(* Logix 5000 project; controller FV vendor 1 type 14 code 217 rev 31.11; software revision 31.00; part 23 of 63 *)
(* tags used below, declared in another part *)
   CheckTimeMask : INT;
   Delphi_Does_Eng_Func : BOOL;
   FR_N255 : INT[265];   // CHECKWORDS
   FR_VB4_AV04 : PlantItem;   // VB4_AV04
   FR_VB4_AV05 : PlantItem;   // VB4_AV05
   FR_VB4_AV06 : PlantItem;   // VB4_AV06
   FR_VB4_AV07 : PlantItem;   // VB4_AV07
   FR_VB4_AV08 : PlantItem;   // VB4_AV08
   FR_VB4_AV09 : PlantItem;   // VB4_AV09
   FR_VB4_AV10 : PlantItem;   // VB4_AV10
   FR_VB4_AV11 : PlantItem;   // VB4_AV11
   FR_VB4_AV12 : PlantItem;   // VB4_AV12
   FR_VB4_AV13 : PlantItem;   // VB4_AV13
   FR_VB4_AV14 : PlantItem;   // VB4_AV14
   FR_VB4_AV15 : PlantItem;   // VB4_AV15
   FR_VB4_AV23 : PlantItem;   // VB4_AV23
   TempChecktime : DINT;
(* FR_Common, continued *)

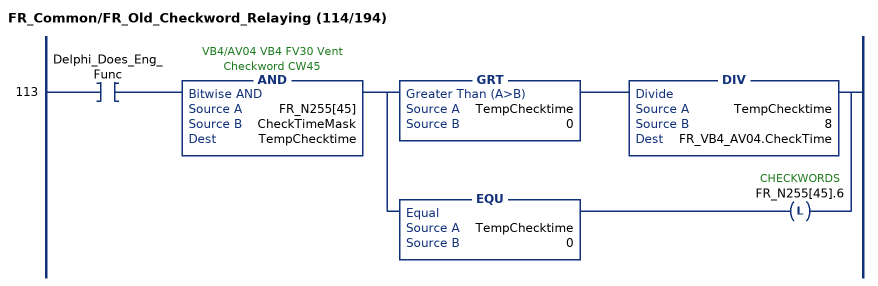
   [picture p418: FR_Common/FR_Old_Checkword_Relaying rungs 113-113]
   113: XIC(Delphi_Does_Eng_Func)AND(FR_N255[45],CheckTimeMask,TempChecktime)[GRT(TempChecktime,0) DIV(TempChecktime,8,FR_VB4_AV04.CheckTime) ,EQU(TempChecktime,0) OTL(FR_N255[45].6) ];
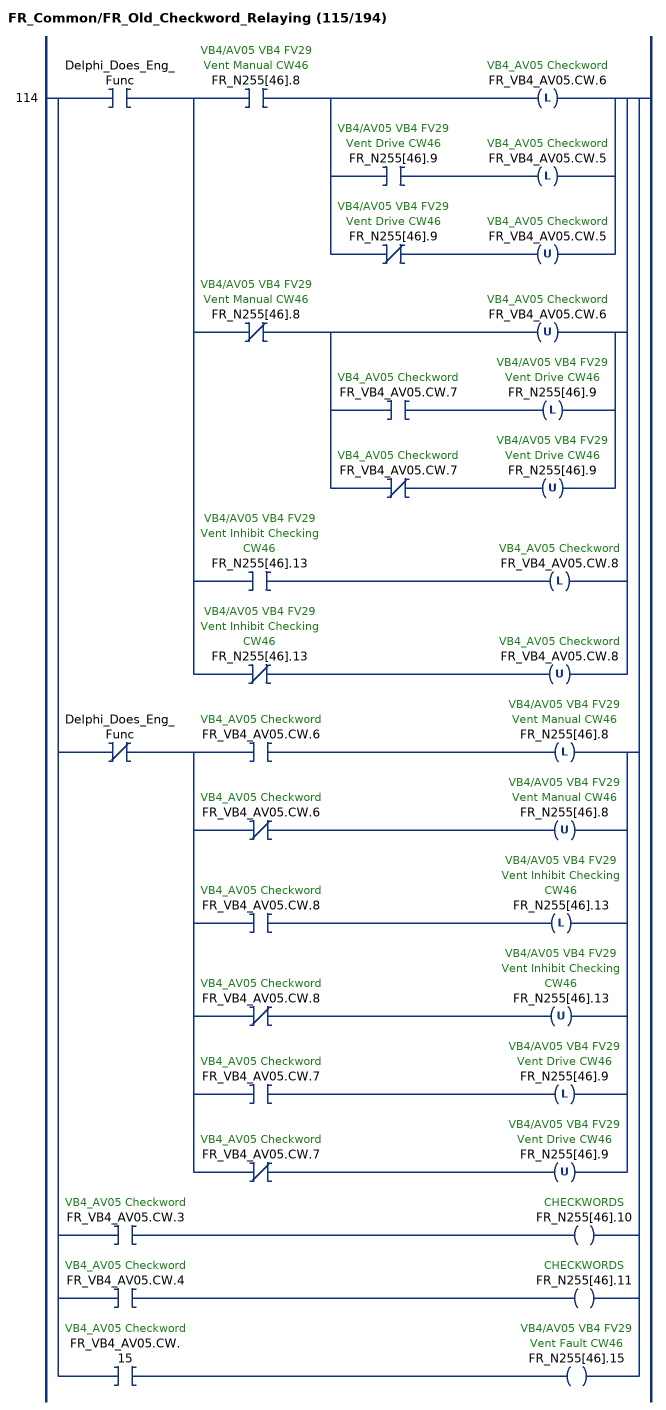
   114: [XIC(Delphi_Does_Eng_Func) [[XIC(FR_N255[46].8) [OTL(FR_VB4_AV05.CW.6) ,XIC(FR_N255[46].9) OTL(FR_VB4_AV05.CW.5) ,XIO(FR_N255[46].9) OTU(FR_VB4_AV05.CW.5) ] ,XIO(FR_N255[46].8) [OTU(FR_VB4_AV05.CW.6) ,[XIC(FR_VB4_AV05.CW.7) OTL(FR_N255[46].9) ,XIO(FR_VB4_AV05.CW.7) OTU(FR_N255[46].9) ] ] ] ,[XIC(FR_N255[46].13) OTL(FR_VB4_AV05.CW.8) ,XIO(FR_N255[46].13) OTU(FR_VB4_AV05.CW.8) ] ] ,XIO(Delphi_Does_Eng_Func) [[XIC(FR_VB4_AV05.CW.6) OTL(FR_N255[46].8) ,XIO(FR_VB4_AV05.CW.6) OTU(FR_N255[46].8) ] ,[XIC(FR_VB4_AV05.CW.8) OTL(FR_N255[46].13) ,XIO(FR_VB4_AV05.CW.8) OTU(FR_N255[46].13) ] ,[XIC(FR_VB4_AV05.CW.7) OTL(FR_N255[46].9) ,XIO(FR_VB4_AV05.CW.7) OTU(FR_N255[46].9) ] ] ,XIC(FR_VB4_AV05.CW.3) OTE(FR_N255[46].10) ,XIC(FR_VB4_AV05.CW.4) OTE(FR_N255[46].11) ,XIC(FR_VB4_AV05.CW.15) OTE(FR_N255[46].15) ];
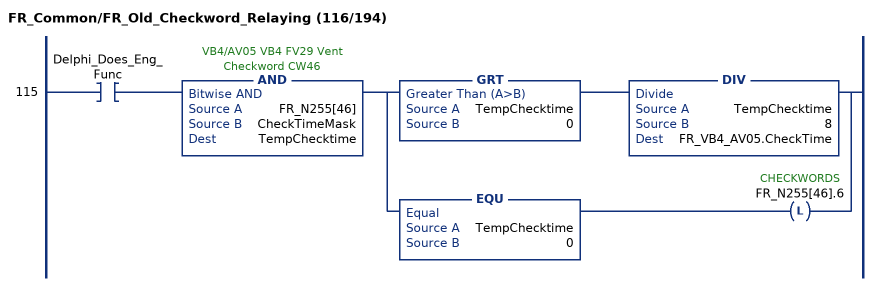
   115: XIC(Delphi_Does_Eng_Func)AND(FR_N255[46],CheckTimeMask,TempChecktime)[GRT(TempChecktime,0) DIV(TempChecktime,8,FR_VB4_AV05.CheckTime) ,EQU(TempChecktime,0) OTL(FR_N255[46].6) ];
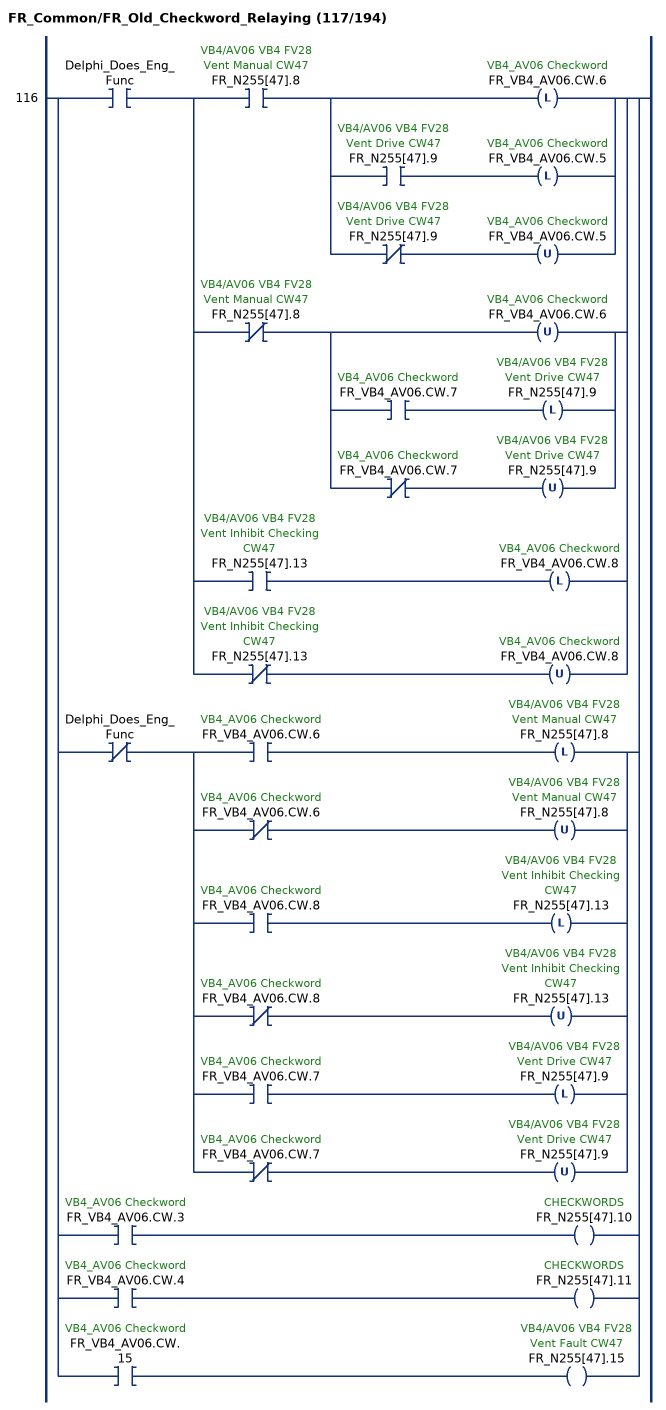
   116: [XIC(Delphi_Does_Eng_Func) [[XIC(FR_N255[47].8) [OTL(FR_VB4_AV06.CW.6) ,XIC(FR_N255[47].9) OTL(FR_VB4_AV06.CW.5) ,XIO(FR_N255[47].9) OTU(FR_VB4_AV06.CW.5) ] ,XIO(FR_N255[47].8) [OTU(FR_VB4_AV06.CW.6) ,[XIC(FR_VB4_AV06.CW.7) OTL(FR_N255[47].9) ,XIO(FR_VB4_AV06.CW.7) OTU(FR_N255[47].9) ] ] ] ,[XIC(FR_N255[47].13) OTL(FR_VB4_AV06.CW.8) ,XIO(FR_N255[47].13) OTU(FR_VB4_AV06.CW.8) ] ] ,XIO(Delphi_Does_Eng_Func) [[XIC(FR_VB4_AV06.CW.6) OTL(FR_N255[47].8) ,XIO(FR_VB4_AV06.CW.6) OTU(FR_N255[47].8) ] ,[XIC(FR_VB4_AV06.CW.8) OTL(FR_N255[47].13) ,XIO(FR_VB4_AV06.CW.8) OTU(FR_N255[47].13) ] ,[XIC(FR_VB4_AV06.CW.7) OTL(FR_N255[47].9) ,XIO(FR_VB4_AV06.CW.7) OTU(FR_N255[47].9) ] ] ,XIC(FR_VB4_AV06.CW.3) OTE(FR_N255[47].10) ,XIC(FR_VB4_AV06.CW.4) OTE(FR_N255[47].11) ,XIC(FR_VB4_AV06.CW.15) OTE(FR_N255[47].15) ];
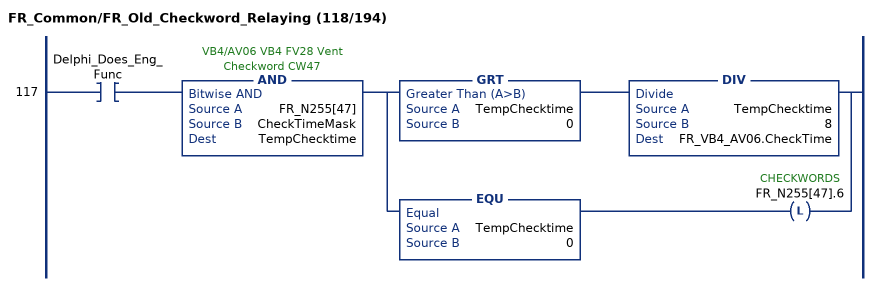
   117: XIC(Delphi_Does_Eng_Func)AND(FR_N255[47],CheckTimeMask,TempChecktime)[GRT(TempChecktime,0) DIV(TempChecktime,8,FR_VB4_AV06.CheckTime) ,EQU(TempChecktime,0) OTL(FR_N255[47].6) ];
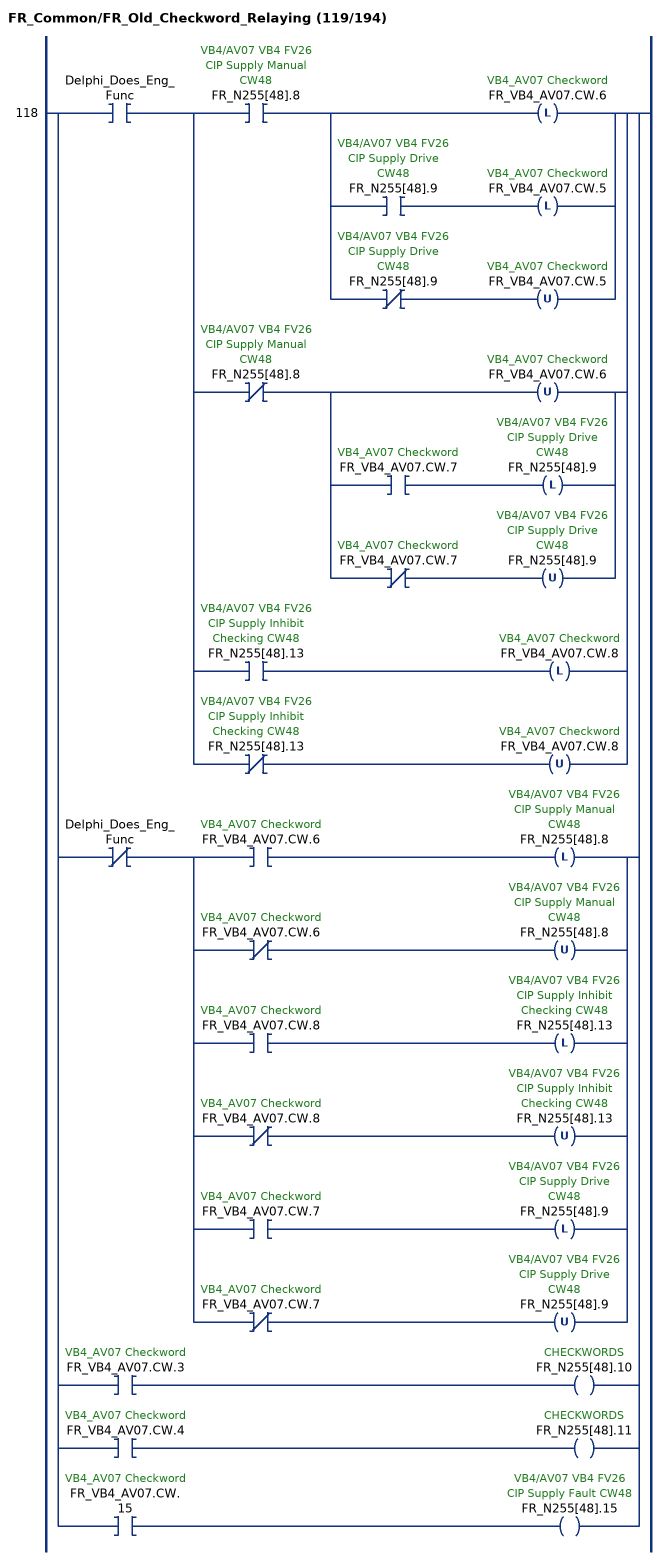
   118: [XIC(Delphi_Does_Eng_Func) [[XIC(FR_N255[48].8) [OTL(FR_VB4_AV07.CW.6) ,XIC(FR_N255[48].9) OTL(FR_VB4_AV07.CW.5) ,XIO(FR_N255[48].9) OTU(FR_VB4_AV07.CW.5) ] ,XIO(FR_N255[48].8) [OTU(FR_VB4_AV07.CW.6) ,[XIC(FR_VB4_AV07.CW.7) OTL(FR_N255[48].9) ,XIO(FR_VB4_AV07.CW.7) OTU(FR_N255[48].9) ] ] ] ,[XIC(FR_N255[48].13) OTL(FR_VB4_AV07.CW.8) ,XIO(FR_N255[48].13) OTU(FR_VB4_AV07.CW.8) ] ] ,XIO(Delphi_Does_Eng_Func) [[XIC(FR_VB4_AV07.CW.6) OTL(FR_N255[48].8) ,XIO(FR_VB4_AV07.CW.6) OTU(FR_N255[48].8) ] ,[XIC(FR_VB4_AV07.CW.8) OTL(FR_N255[48].13) ,XIO(FR_VB4_AV07.CW.8) OTU(FR_N255[48].13) ] ,[XIC(FR_VB4_AV07.CW.7) OTL(FR_N255[48].9) ,XIO(FR_VB4_AV07.CW.7) OTU(FR_N255[48].9) ] ] ,XIC(FR_VB4_AV07.CW.3) OTE(FR_N255[48].10) ,XIC(FR_VB4_AV07.CW.4) OTE(FR_N255[48].11) ,XIC(FR_VB4_AV07.CW.15) OTE(FR_N255[48].15) ];
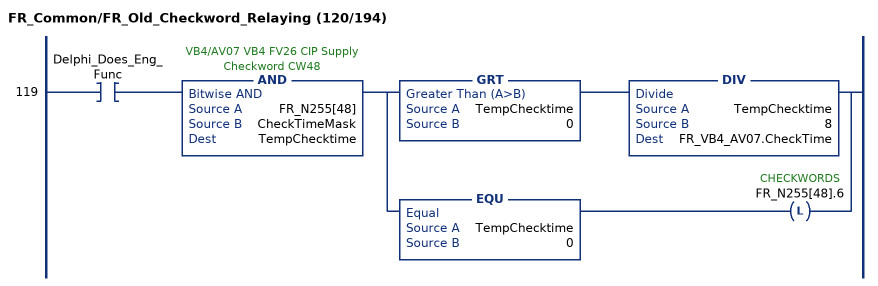
   119: XIC(Delphi_Does_Eng_Func)AND(FR_N255[48],CheckTimeMask,TempChecktime)[GRT(TempChecktime,0) DIV(TempChecktime,8,FR_VB4_AV07.CheckTime) ,EQU(TempChecktime,0) OTL(FR_N255[48].6) ];
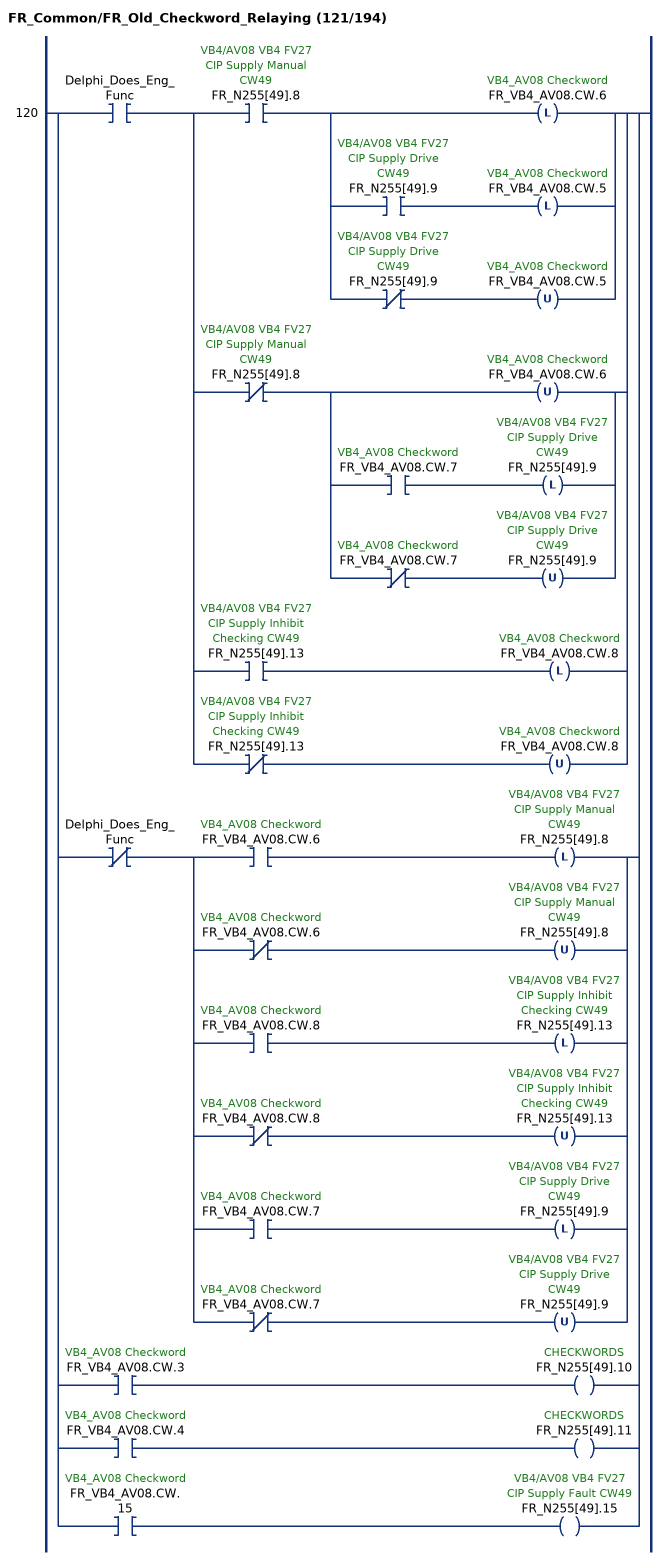
   120: [XIC(Delphi_Does_Eng_Func) [[XIC(FR_N255[49].8) [OTL(FR_VB4_AV08.CW.6) ,XIC(FR_N255[49].9) OTL(FR_VB4_AV08.CW.5) ,XIO(FR_N255[49].9) OTU(FR_VB4_AV08.CW.5) ] ,XIO(FR_N255[49].8) [OTU(FR_VB4_AV08.CW.6) ,[XIC(FR_VB4_AV08.CW.7) OTL(FR_N255[49].9) ,XIO(FR_VB4_AV08.CW.7) OTU(FR_N255[49].9) ] ] ] ,[XIC(FR_N255[49].13) OTL(FR_VB4_AV08.CW.8) ,XIO(FR_N255[49].13) OTU(FR_VB4_AV08.CW.8) ] ] ,XIO(Delphi_Does_Eng_Func) [[XIC(FR_VB4_AV08.CW.6) OTL(FR_N255[49].8) ,XIO(FR_VB4_AV08.CW.6) OTU(FR_N255[49].8) ] ,[XIC(FR_VB4_AV08.CW.8) OTL(FR_N255[49].13) ,XIO(FR_VB4_AV08.CW.8) OTU(FR_N255[49].13) ] ,[XIC(FR_VB4_AV08.CW.7) OTL(FR_N255[49].9) ,XIO(FR_VB4_AV08.CW.7) OTU(FR_N255[49].9) ] ] ,XIC(FR_VB4_AV08.CW.3) OTE(FR_N255[49].10) ,XIC(FR_VB4_AV08.CW.4) OTE(FR_N255[49].11) ,XIC(FR_VB4_AV08.CW.15) OTE(FR_N255[49].15) ];
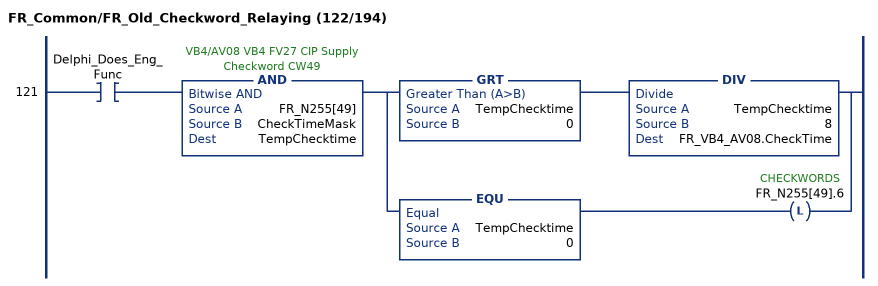
   121: XIC(Delphi_Does_Eng_Func)AND(FR_N255[49],CheckTimeMask,TempChecktime)[GRT(TempChecktime,0) DIV(TempChecktime,8,FR_VB4_AV08.CheckTime) ,EQU(TempChecktime,0) OTL(FR_N255[49].6) ];
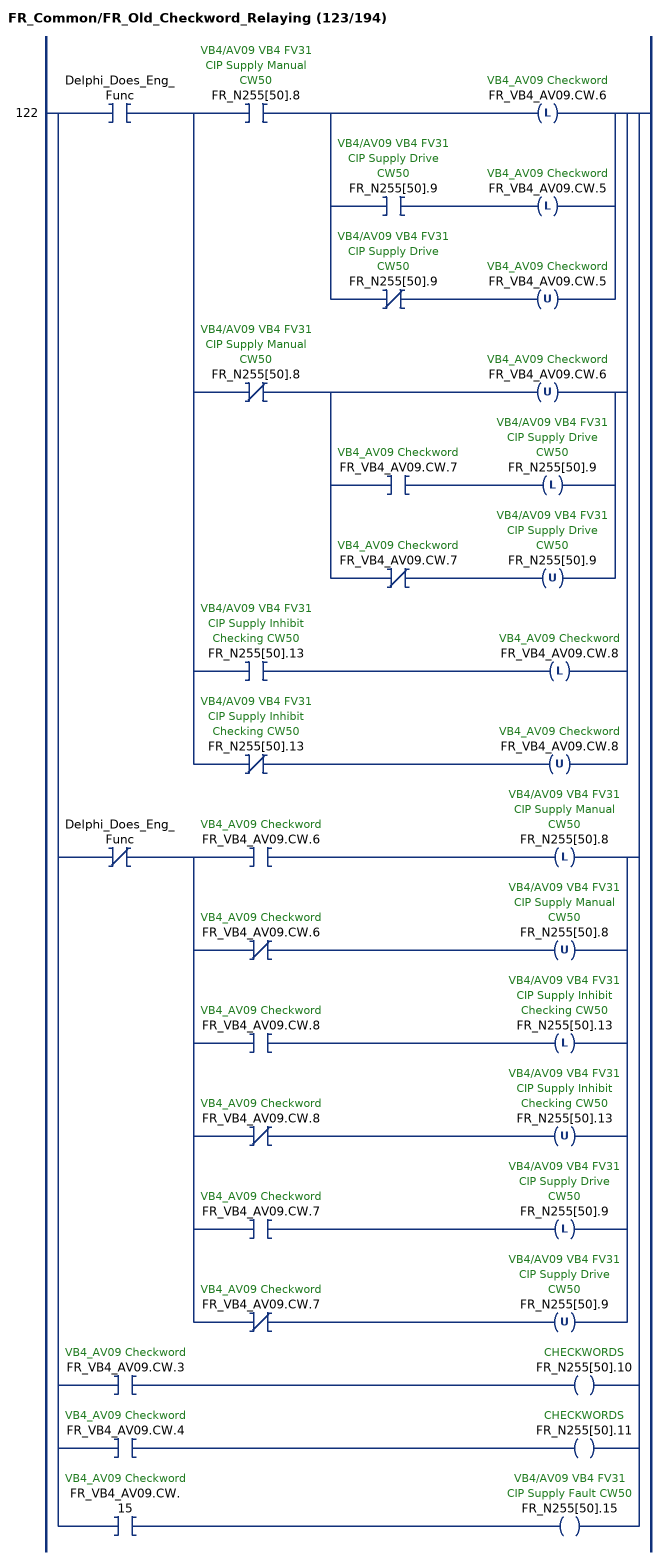
   122: [XIC(Delphi_Does_Eng_Func) [[XIC(FR_N255[50].8) [OTL(FR_VB4_AV09.CW.6) ,XIC(FR_N255[50].9) OTL(FR_VB4_AV09.CW.5) ,XIO(FR_N255[50].9) OTU(FR_VB4_AV09.CW.5) ] ,XIO(FR_N255[50].8) [OTU(FR_VB4_AV09.CW.6) ,[XIC(FR_VB4_AV09.CW.7) OTL(FR_N255[50].9) ,XIO(FR_VB4_AV09.CW.7) OTU(FR_N255[50].9) ] ] ] ,[XIC(FR_N255[50].13) OTL(FR_VB4_AV09.CW.8) ,XIO(FR_N255[50].13) OTU(FR_VB4_AV09.CW.8) ] ] ,XIO(Delphi_Does_Eng_Func) [[XIC(FR_VB4_AV09.CW.6) OTL(FR_N255[50].8) ,XIO(FR_VB4_AV09.CW.6) OTU(FR_N255[50].8) ] ,[XIC(FR_VB4_AV09.CW.8) OTL(FR_N255[50].13) ,XIO(FR_VB4_AV09.CW.8) OTU(FR_N255[50].13) ] ,[XIC(FR_VB4_AV09.CW.7) OTL(FR_N255[50].9) ,XIO(FR_VB4_AV09.CW.7) OTU(FR_N255[50].9) ] ] ,XIC(FR_VB4_AV09.CW.3) OTE(FR_N255[50].10) ,XIC(FR_VB4_AV09.CW.4) OTE(FR_N255[50].11) ,XIC(FR_VB4_AV09.CW.15) OTE(FR_N255[50].15) ];
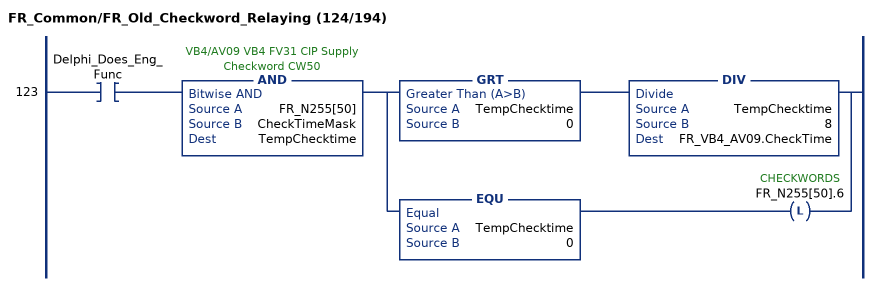
   123: XIC(Delphi_Does_Eng_Func)AND(FR_N255[50],CheckTimeMask,TempChecktime)[GRT(TempChecktime,0) DIV(TempChecktime,8,FR_VB4_AV09.CheckTime) ,EQU(TempChecktime,0) OTL(FR_N255[50].6) ];
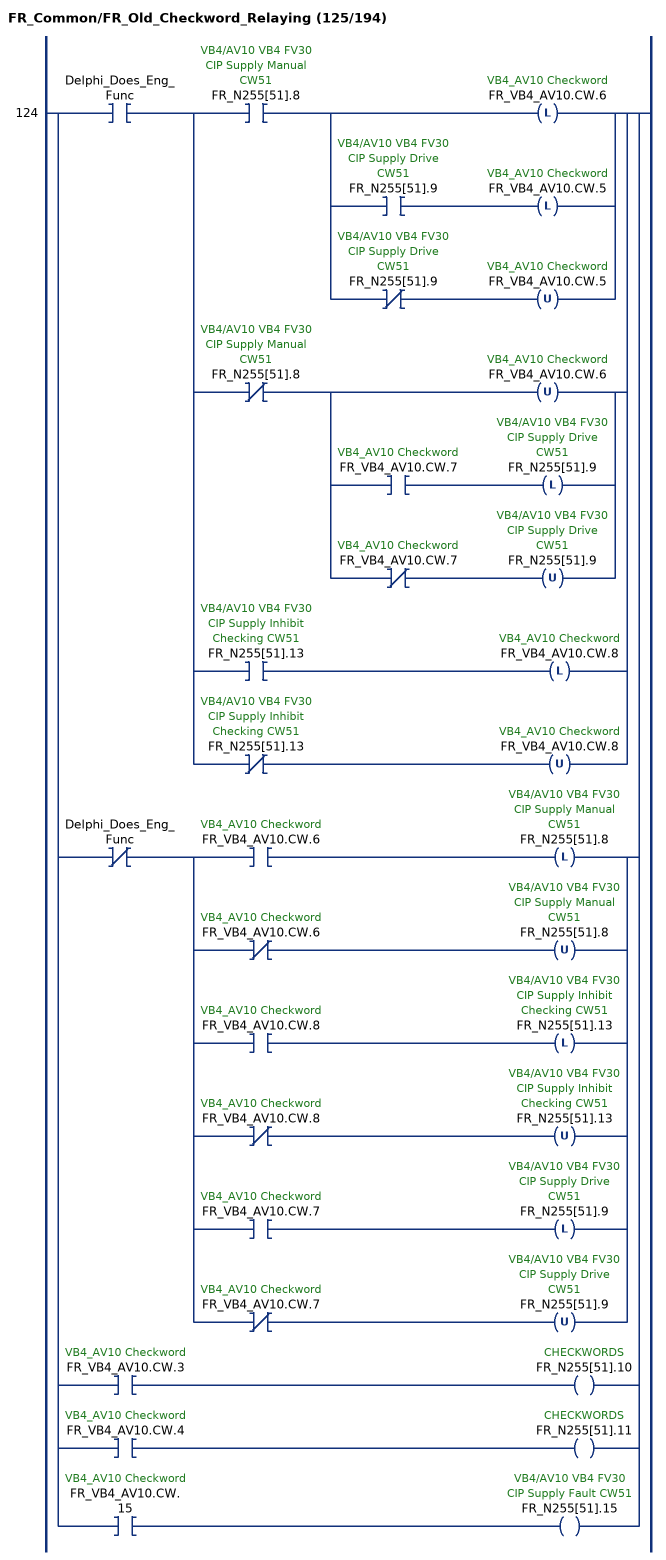
   124: [XIC(Delphi_Does_Eng_Func) [[XIC(FR_N255[51].8) [OTL(FR_VB4_AV10.CW.6) ,XIC(FR_N255[51].9) OTL(FR_VB4_AV10.CW.5) ,XIO(FR_N255[51].9) OTU(FR_VB4_AV10.CW.5) ] ,XIO(FR_N255[51].8) [OTU(FR_VB4_AV10.CW.6) ,[XIC(FR_VB4_AV10.CW.7) OTL(FR_N255[51].9) ,XIO(FR_VB4_AV10.CW.7) OTU(FR_N255[51].9) ] ] ] ,[XIC(FR_N255[51].13) OTL(FR_VB4_AV10.CW.8) ,XIO(FR_N255[51].13) OTU(FR_VB4_AV10.CW.8) ] ] ,XIO(Delphi_Does_Eng_Func) [[XIC(FR_VB4_AV10.CW.6) OTL(FR_N255[51].8) ,XIO(FR_VB4_AV10.CW.6) OTU(FR_N255[51].8) ] ,[XIC(FR_VB4_AV10.CW.8) OTL(FR_N255[51].13) ,XIO(FR_VB4_AV10.CW.8) OTU(FR_N255[51].13) ] ,[XIC(FR_VB4_AV10.CW.7) OTL(FR_N255[51].9) ,XIO(FR_VB4_AV10.CW.7) OTU(FR_N255[51].9) ] ] ,XIC(FR_VB4_AV10.CW.3) OTE(FR_N255[51].10) ,XIC(FR_VB4_AV10.CW.4) OTE(FR_N255[51].11) ,XIC(FR_VB4_AV10.CW.15) OTE(FR_N255[51].15) ];
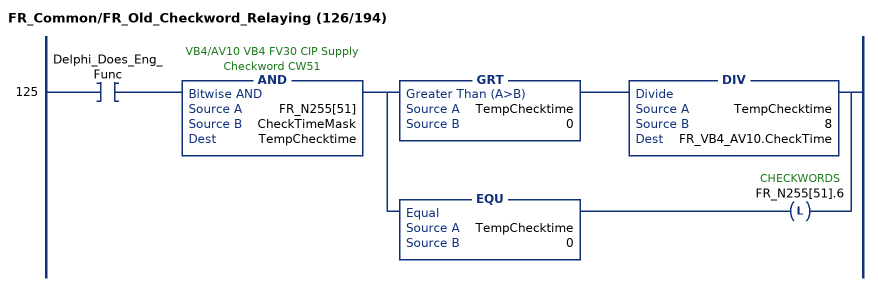
   125: XIC(Delphi_Does_Eng_Func)AND(FR_N255[51],CheckTimeMask,TempChecktime)[GRT(TempChecktime,0) DIV(TempChecktime,8,FR_VB4_AV10.CheckTime) ,EQU(TempChecktime,0) OTL(FR_N255[51].6) ];
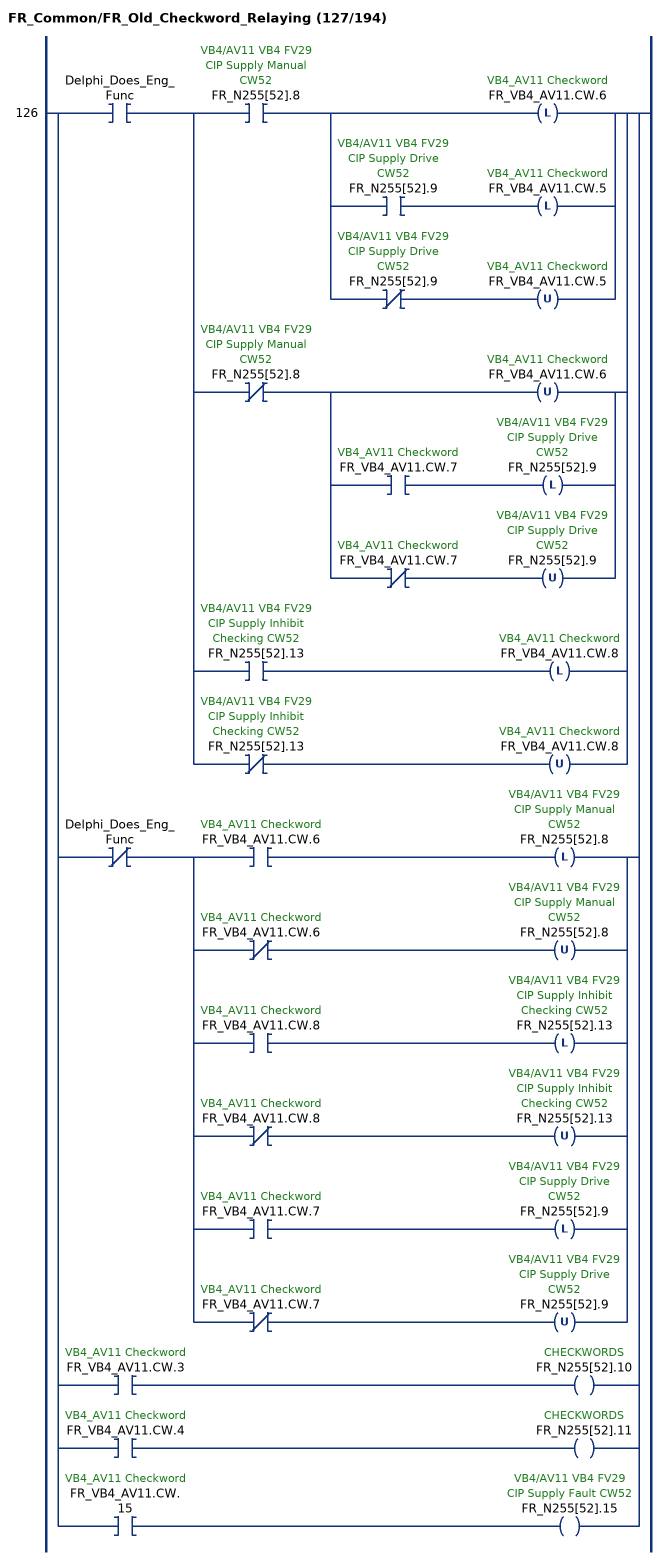
   126: [XIC(Delphi_Does_Eng_Func) [[XIC(FR_N255[52].8) [OTL(FR_VB4_AV11.CW.6) ,XIC(FR_N255[52].9) OTL(FR_VB4_AV11.CW.5) ,XIO(FR_N255[52].9) OTU(FR_VB4_AV11.CW.5) ] ,XIO(FR_N255[52].8) [OTU(FR_VB4_AV11.CW.6) ,[XIC(FR_VB4_AV11.CW.7) OTL(FR_N255[52].9) ,XIO(FR_VB4_AV11.CW.7) OTU(FR_N255[52].9) ] ] ] ,[XIC(FR_N255[52].13) OTL(FR_VB4_AV11.CW.8) ,XIO(FR_N255[52].13) OTU(FR_VB4_AV11.CW.8) ] ] ,XIO(Delphi_Does_Eng_Func) [[XIC(FR_VB4_AV11.CW.6) OTL(FR_N255[52].8) ,XIO(FR_VB4_AV11.CW.6) OTU(FR_N255[52].8) ] ,[XIC(FR_VB4_AV11.CW.8) OTL(FR_N255[52].13) ,XIO(FR_VB4_AV11.CW.8) OTU(FR_N255[52].13) ] ,[XIC(FR_VB4_AV11.CW.7) OTL(FR_N255[52].9) ,XIO(FR_VB4_AV11.CW.7) OTU(FR_N255[52].9) ] ] ,XIC(FR_VB4_AV11.CW.3) OTE(FR_N255[52].10) ,XIC(FR_VB4_AV11.CW.4) OTE(FR_N255[52].11) ,XIC(FR_VB4_AV11.CW.15) OTE(FR_N255[52].15) ];
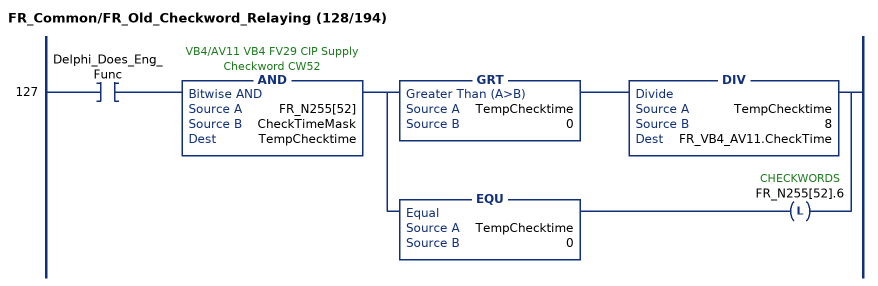
   127: XIC(Delphi_Does_Eng_Func)AND(FR_N255[52],CheckTimeMask,TempChecktime)[GRT(TempChecktime,0) DIV(TempChecktime,8,FR_VB4_AV11.CheckTime) ,EQU(TempChecktime,0) OTL(FR_N255[52].6) ];
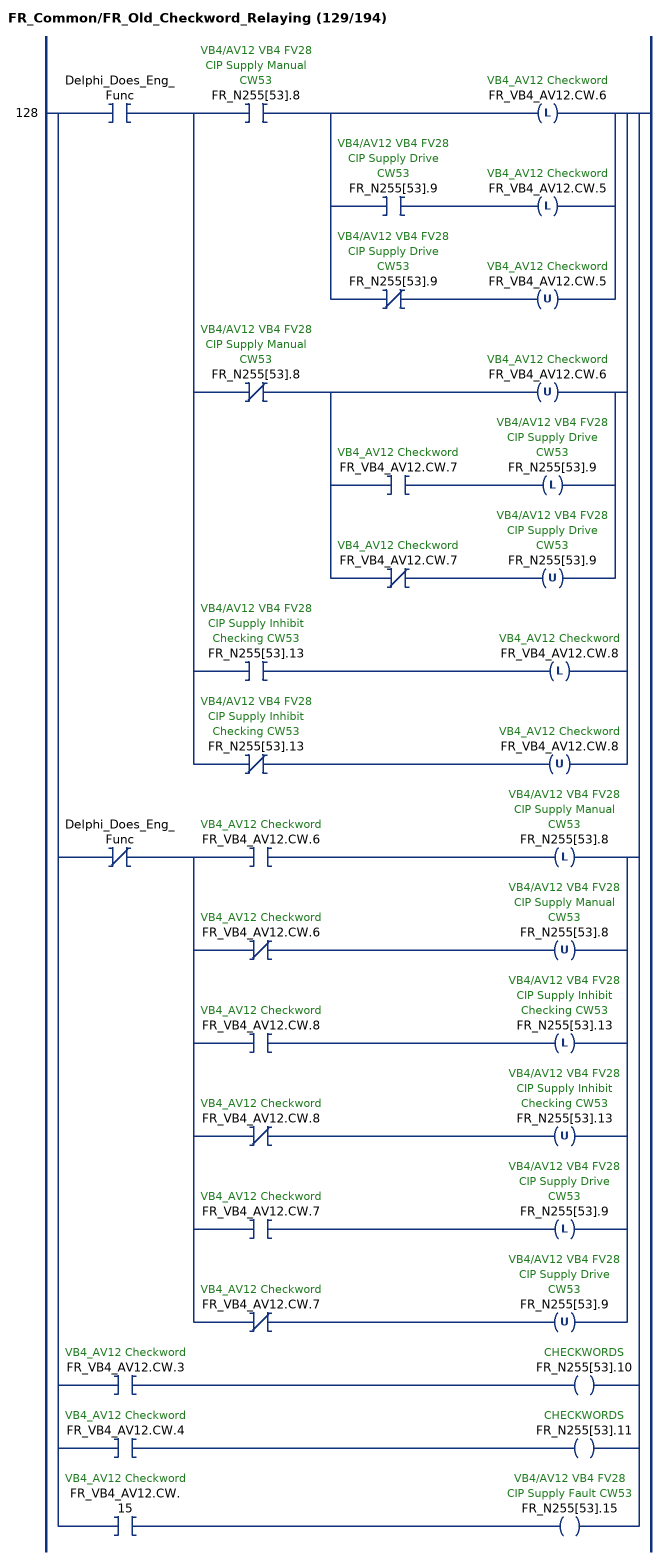
   128: [XIC(Delphi_Does_Eng_Func) [[XIC(FR_N255[53].8) [OTL(FR_VB4_AV12.CW.6) ,XIC(FR_N255[53].9) OTL(FR_VB4_AV12.CW.5) ,XIO(FR_N255[53].9) OTU(FR_VB4_AV12.CW.5) ] ,XIO(FR_N255[53].8) [OTU(FR_VB4_AV12.CW.6) ,[XIC(FR_VB4_AV12.CW.7) OTL(FR_N255[53].9) ,XIO(FR_VB4_AV12.CW.7) OTU(FR_N255[53].9) ] ] ] ,[XIC(FR_N255[53].13) OTL(FR_VB4_AV12.CW.8) ,XIO(FR_N255[53].13) OTU(FR_VB4_AV12.CW.8) ] ] ,XIO(Delphi_Does_Eng_Func) [[XIC(FR_VB4_AV12.CW.6) OTL(FR_N255[53].8) ,XIO(FR_VB4_AV12.CW.6) OTU(FR_N255[53].8) ] ,[XIC(FR_VB4_AV12.CW.8) OTL(FR_N255[53].13) ,XIO(FR_VB4_AV12.CW.8) OTU(FR_N255[53].13) ] ,[XIC(FR_VB4_AV12.CW.7) OTL(FR_N255[53].9) ,XIO(FR_VB4_AV12.CW.7) OTU(FR_N255[53].9) ] ] ,XIC(FR_VB4_AV12.CW.3) OTE(FR_N255[53].10) ,XIC(FR_VB4_AV12.CW.4) OTE(FR_N255[53].11) ,XIC(FR_VB4_AV12.CW.15) OTE(FR_N255[53].15) ];
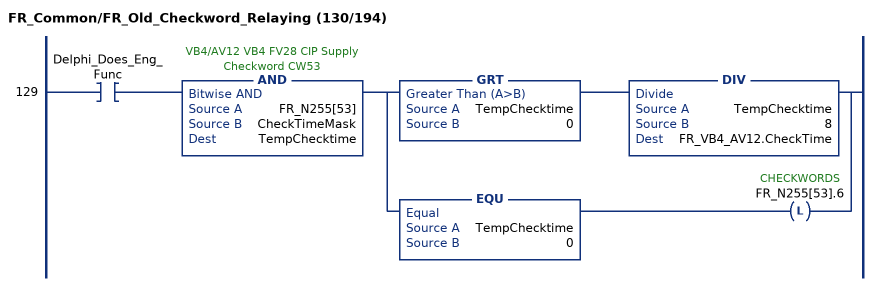
   129: XIC(Delphi_Does_Eng_Func)AND(FR_N255[53],CheckTimeMask,TempChecktime)[GRT(TempChecktime,0) DIV(TempChecktime,8,FR_VB4_AV12.CheckTime) ,EQU(TempChecktime,0) OTL(FR_N255[53].6) ];
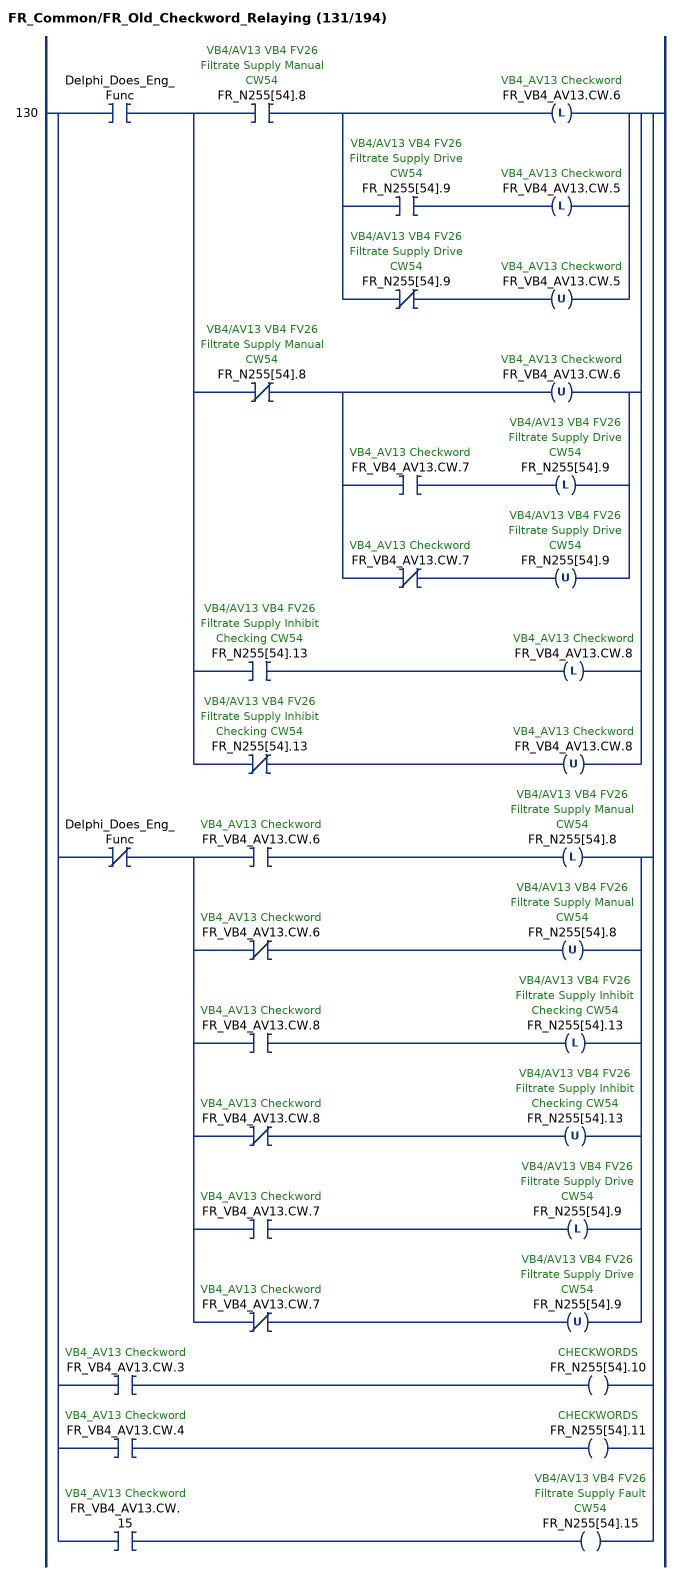
   130: [XIC(Delphi_Does_Eng_Func) [[XIC(FR_N255[54].8) [OTL(FR_VB4_AV13.CW.6) ,XIC(FR_N255[54].9) OTL(FR_VB4_AV13.CW.5) ,XIO(FR_N255[54].9) OTU(FR_VB4_AV13.CW.5) ] ,XIO(FR_N255[54].8) [OTU(FR_VB4_AV13.CW.6) ,[XIC(FR_VB4_AV13.CW.7) OTL(FR_N255[54].9) ,XIO(FR_VB4_AV13.CW.7) OTU(FR_N255[54].9) ] ] ] ,[XIC(FR_N255[54].13) OTL(FR_VB4_AV13.CW.8) ,XIO(FR_N255[54].13) OTU(FR_VB4_AV13.CW.8) ] ] ,XIO(Delphi_Does_Eng_Func) [[XIC(FR_VB4_AV13.CW.6) OTL(FR_N255[54].8) ,XIO(FR_VB4_AV13.CW.6) OTU(FR_N255[54].8) ] ,[XIC(FR_VB4_AV13.CW.8) OTL(FR_N255[54].13) ,XIO(FR_VB4_AV13.CW.8) OTU(FR_N255[54].13) ] ,[XIC(FR_VB4_AV13.CW.7) OTL(FR_N255[54].9) ,XIO(FR_VB4_AV13.CW.7) OTU(FR_N255[54].9) ] ] ,XIC(FR_VB4_AV13.CW.3) OTE(FR_N255[54].10) ,XIC(FR_VB4_AV13.CW.4) OTE(FR_N255[54].11) ,XIC(FR_VB4_AV13.CW.15) OTE(FR_N255[54].15) ];
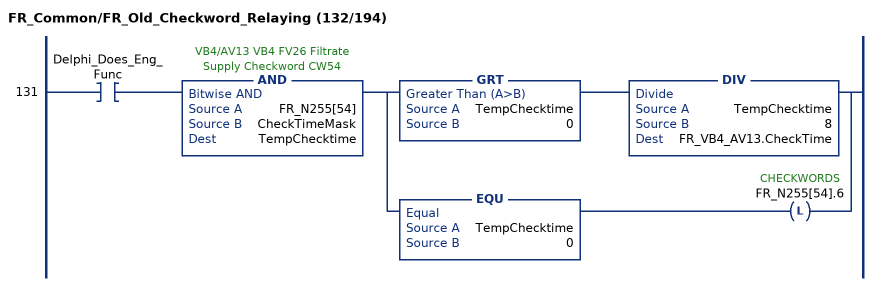
   131: XIC(Delphi_Does_Eng_Func)AND(FR_N255[54],CheckTimeMask,TempChecktime)[GRT(TempChecktime,0) DIV(TempChecktime,8,FR_VB4_AV13.CheckTime) ,EQU(TempChecktime,0) OTL(FR_N255[54].6) ];
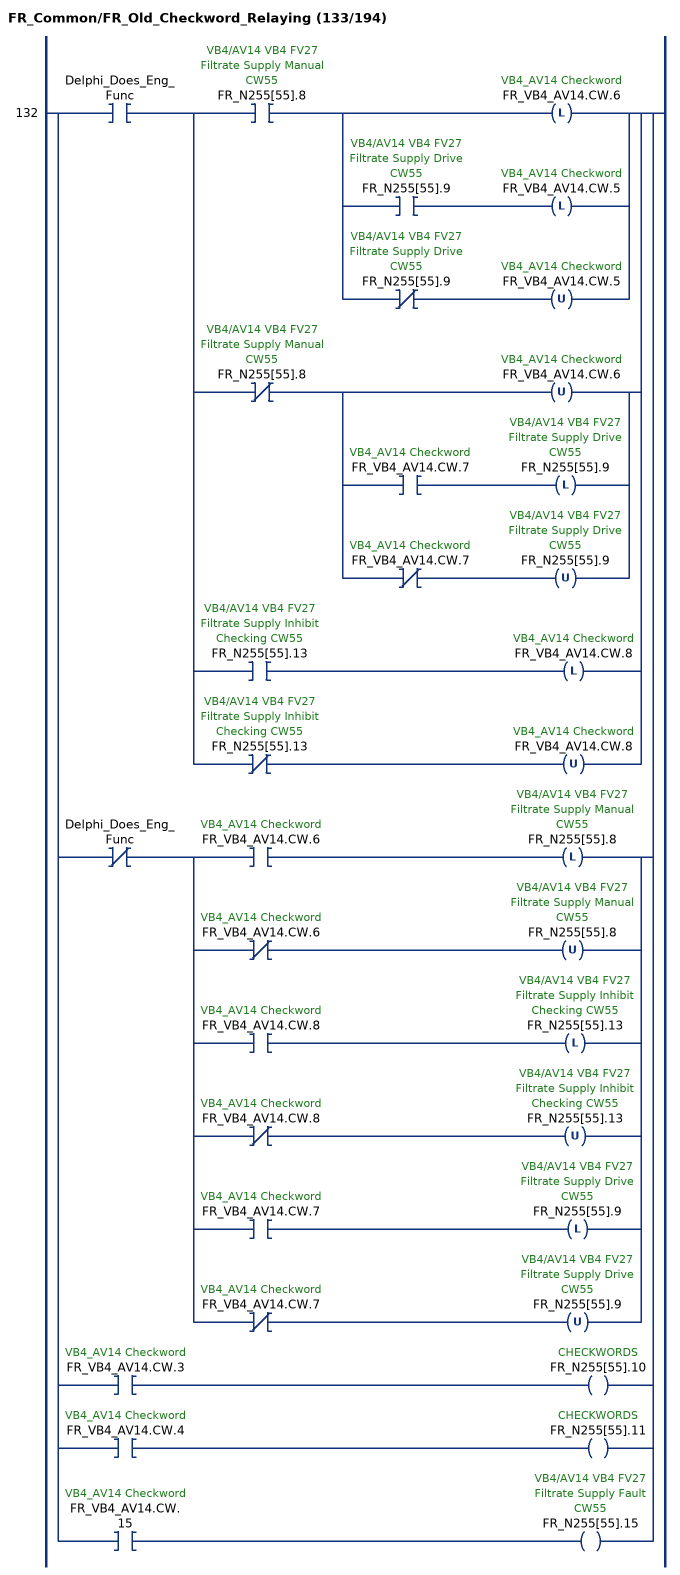
   132: [XIC(Delphi_Does_Eng_Func) [[XIC(FR_N255[55].8) [OTL(FR_VB4_AV14.CW.6) ,XIC(FR_N255[55].9) OTL(FR_VB4_AV14.CW.5) ,XIO(FR_N255[55].9) OTU(FR_VB4_AV14.CW.5) ] ,XIO(FR_N255[55].8) [OTU(FR_VB4_AV14.CW.6) ,[XIC(FR_VB4_AV14.CW.7) OTL(FR_N255[55].9) ,XIO(FR_VB4_AV14.CW.7) OTU(FR_N255[55].9) ] ] ] ,[XIC(FR_N255[55].13) OTL(FR_VB4_AV14.CW.8) ,XIO(FR_N255[55].13) OTU(FR_VB4_AV14.CW.8) ] ] ,XIO(Delphi_Does_Eng_Func) [[XIC(FR_VB4_AV14.CW.6) OTL(FR_N255[55].8) ,XIO(FR_VB4_AV14.CW.6) OTU(FR_N255[55].8) ] ,[XIC(FR_VB4_AV14.CW.8) OTL(FR_N255[55].13) ,XIO(FR_VB4_AV14.CW.8) OTU(FR_N255[55].13) ] ,[XIC(FR_VB4_AV14.CW.7) OTL(FR_N255[55].9) ,XIO(FR_VB4_AV14.CW.7) OTU(FR_N255[55].9) ] ] ,XIC(FR_VB4_AV14.CW.3) OTE(FR_N255[55].10) ,XIC(FR_VB4_AV14.CW.4) OTE(FR_N255[55].11) ,XIC(FR_VB4_AV14.CW.15) OTE(FR_N255[55].15) ];
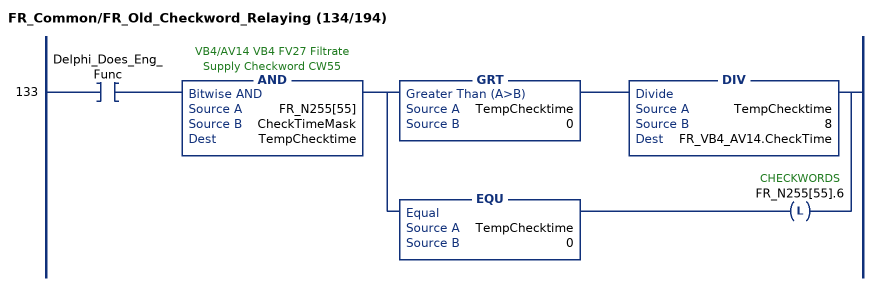
   133: XIC(Delphi_Does_Eng_Func)AND(FR_N255[55],CheckTimeMask,TempChecktime)[GRT(TempChecktime,0) DIV(TempChecktime,8,FR_VB4_AV14.CheckTime) ,EQU(TempChecktime,0) OTL(FR_N255[55].6) ];
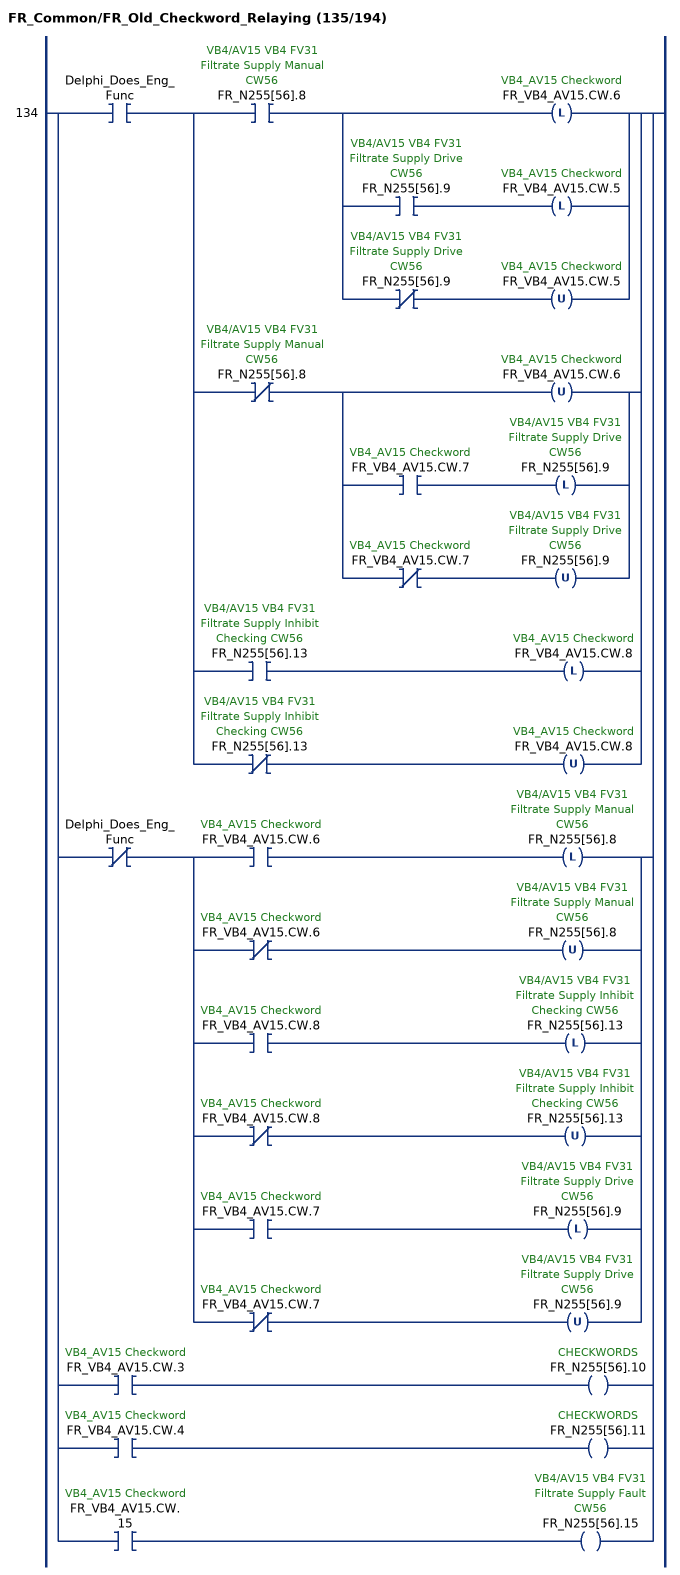
   134: [XIC(Delphi_Does_Eng_Func) [[XIC(FR_N255[56].8) [OTL(FR_VB4_AV15.CW.6) ,XIC(FR_N255[56].9) OTL(FR_VB4_AV15.CW.5) ,XIO(FR_N255[56].9) OTU(FR_VB4_AV15.CW.5) ] ,XIO(FR_N255[56].8) [OTU(FR_VB4_AV15.CW.6) ,[XIC(FR_VB4_AV15.CW.7) OTL(FR_N255[56].9) ,XIO(FR_VB4_AV15.CW.7) OTU(FR_N255[56].9) ] ] ] ,[XIC(FR_N255[56].13) OTL(FR_VB4_AV15.CW.8) ,XIO(FR_N255[56].13) OTU(FR_VB4_AV15.CW.8) ] ] ,XIO(Delphi_Does_Eng_Func) [[XIC(FR_VB4_AV15.CW.6) OTL(FR_N255[56].8) ,XIO(FR_VB4_AV15.CW.6) OTU(FR_N255[56].8) ] ,[XIC(FR_VB4_AV15.CW.8) OTL(FR_N255[56].13) ,XIO(FR_VB4_AV15.CW.8) OTU(FR_N255[56].13) ] ,[XIC(FR_VB4_AV15.CW.7) OTL(FR_N255[56].9) ,XIO(FR_VB4_AV15.CW.7) OTU(FR_N255[56].9) ] ] ,XIC(FR_VB4_AV15.CW.3) OTE(FR_N255[56].10) ,XIC(FR_VB4_AV15.CW.4) OTE(FR_N255[56].11) ,XIC(FR_VB4_AV15.CW.15) OTE(FR_N255[56].15) ];
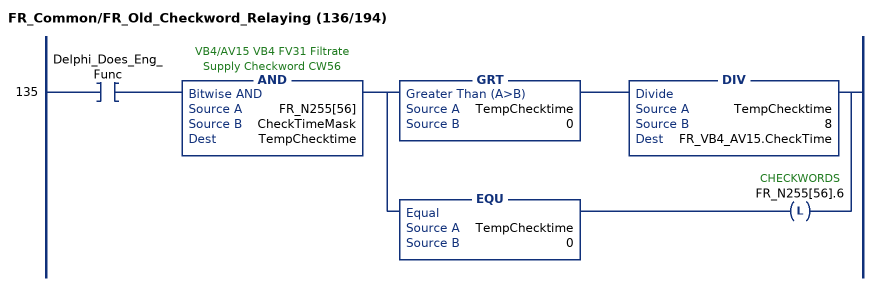
   135: XIC(Delphi_Does_Eng_Func)AND(FR_N255[56],CheckTimeMask,TempChecktime)[GRT(TempChecktime,0) DIV(TempChecktime,8,FR_VB4_AV15.CheckTime) ,EQU(TempChecktime,0) OTL(FR_N255[56].6) ];
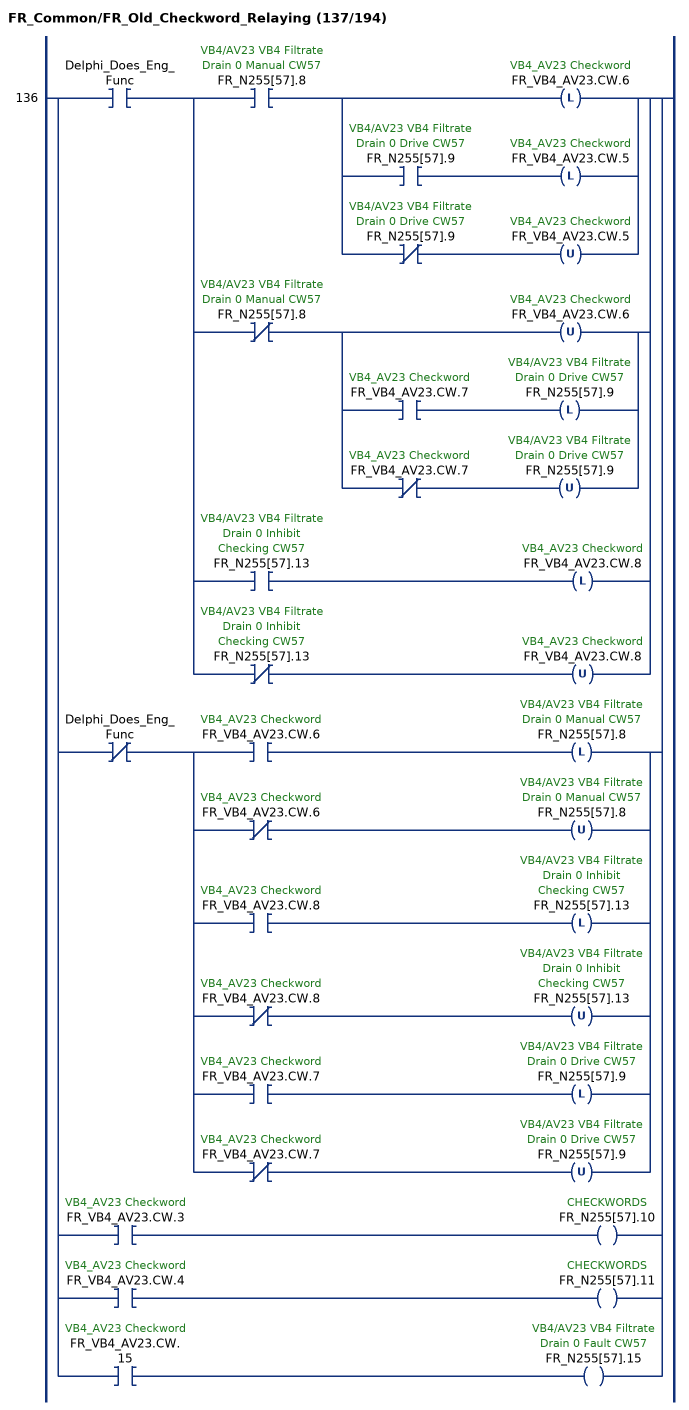
   136: [XIC(Delphi_Does_Eng_Func) [[XIC(FR_N255[57].8) [OTL(FR_VB4_AV23.CW.6) ,XIC(FR_N255[57].9) OTL(FR_VB4_AV23.CW.5) ,XIO(FR_N255[57].9) OTU(FR_VB4_AV23.CW.5) ] ,XIO(FR_N255[57].8) [OTU(FR_VB4_AV23.CW.6) ,[XIC(FR_VB4_AV23.CW.7) OTL(FR_N255[57].9) ,XIO(FR_VB4_AV23.CW.7) OTU(FR_N255[57].9) ] ] ] ,[XIC(FR_N255[57].13) OTL(FR_VB4_AV23.CW.8) ,XIO(FR_N255[57].13) OTU(FR_VB4_AV23.CW.8) ] ] ,XIO(Delphi_Does_Eng_Func) [[XIC(FR_VB4_AV23.CW.6) OTL(FR_N255[57].8) ,XIO(FR_VB4_AV23.CW.6) OTU(FR_N255[57].8) ] ,[XIC(FR_VB4_AV23.CW.8) OTL(FR_N255[57].13) ,XIO(FR_VB4_AV23.CW.8) OTU(FR_N255[57].13) ] ,[XIC(FR_VB4_AV23.CW.7) OTL(FR_N255[57].9) ,XIO(FR_VB4_AV23.CW.7) OTU(FR_N255[57].9) ] ] ,XIC(FR_VB4_AV23.CW.3) OTE(FR_N255[57].10) ,XIC(FR_VB4_AV23.CW.4) OTE(FR_N255[57].11) ,XIC(FR_VB4_AV23.CW.15) OTE(FR_N255[57].15) ];
